
         L     0;
         T     #STC_tPROP.iSyncState;
         L     3;
         T     #OUT_iRetVal;
         BEU;

   e006: A     #STC_tW_MngSysReg.tST.xDone;
         JCN   s006;

         L     6;
         T     #STC_tPROP.iSyncState;

         CALL  FILL
         ( BVAL    := #TMP_dZero,
           RET_VAL := #TMP_iAuxRetVal,
           BLK     := #STC_tW_MngSysReg
         );
         JU    out;
   s006: NOP   0;
END_REGION

REGION Network 9 (STL): RESET "PING" (BIT 1) IN STW1 OF CU
         L     #STC_tPROP.iSyncState;
         L     6;
         ==I;
         JCN   s007;

         SET;
         R     #STC_tPZD_CU.tW.tSTW1.x1;

         L     7;
         T     #STC_tPROP.iSyncState;
         JU    out;
   s007: NOP   0;
END_REGION

REGION Network 10 (STL): SET DONE
         L     #STC_tPROP.iSyncState;
         L     7;
         ==I;
         JCN   s008;

         S     #OUT_xDone;

         L     W#16#0;
         T     #STC_tPROP.iSyncState;

   s008: NOP   0;
END_REGION

REGION Network 11 (STL): Copy Output
   out:  L     #STC_tSYS_DATA.iIOAddress_CU;
         SLW   3;
         T     #TMP_dIO_Pointer;

         L;
         +     48;
         T     #TMP_dPZD_Pointer;

         L     DIW[ #TMP_dPZD_Pointer];
         L     W#16#2;
         AW;
         L     QW[ #TMP_dIO_Pointer];
         OW;
         T     QW[ #TMP_dIO_Pointer];

         BEU;
END_REGION

REGION Network 12 (STL): CU Address wrong
   NWCU: SET;
         S     #OUT_xError;

         L     4;
         T     #OUT_iRetVal;
END_REGION
END_FUNCTION_BLOCK

// folder: 03_Programs_Logics/MCC1201/30_InterfaceEmergencyCutting

FUNCTION_BLOCK "FB_IO_EmergencyCuttingBridge"   // FB28, LAD
{ S7_Optimized_Access := 'TRUE' }
VERSION : 0.1
   VAR_INPUT
      IN_xCycleON : Bool;   // Cycle ON
      IN_xCycleONDel : Bool;   // Delayed cycle ON signal
      IN_xResetAlarms : Bool;   // Reset alarms
      IN_xFaultsEnabled : Bool;   // Faults enabled
      IN_xMachineReady : Bool;   // Machine ready
      IN_xStartCutCycle : Bool;   // StartCutCycle
      IN_xStartCutForBreak : Bool;
      IN_xProtection : Bool;   // EM Xcut protection
      IN_dConvSpeed : DInt;
      IN_xSimulationActive : Bool;
   END_VAR
   VAR_OUTPUT
      OUT_xStartCutCycle : Bool;
      OUT_xSpare : Bool;
      OUT_xSnap : Bool;
      OUT_xAccelaration : Bool;
   END_VAR
   VAR
      ST_xMachineAnomaly : Bool;   // Machine anomaly
      ST_xStoppingFaults : Bool;   // Stopping fault
      ST_xFaults : Bool;   // Fault
      ST_xWarnings : Bool;   // Warnings
      ST_xConditionOkStopCycle : Bool;   // Condition ok stop cycle
      ST_xOutputEnable : Bool;   // Output enable
      ST_xStartcut : Bool;   // Start Cut
      ST_xStartCutForTrak : Bool;
      ST_xRiseAfterDescence : Bool;
      ST_TrackingOnZone_0 : Bool;   // ST_Tracking On Zone0 (0-500)
      ST_TrackingOnZone_1 : Bool;   // ST_Tracking On Zone0 (500-1000)
      ST_TrackingOnZone_2 : Bool;   // ST_Tracking On Zone0 (1000-1500)
      ST_TrackingOnZone_3 : Bool;   // ST_Tracking On Zone0 (1500-2000)
      ST_TrackingOnZone_4 : Bool;   // ST_Tracking On Zone0 (2500-3000)
      ST_TrackingOnZone_5 : Bool;   // ST_Tracking On Zone0 (3500-4000)
      ST_TrackingOnZone_6 : Bool;   // ST_Tracking On Zone0 (3500-4000)
      Os_Ready : Bool;
      Os_Readys : Bool;
      Os_StartCut : Bool;
      OSR_CyclecuttingON : Bool;
      OUTPUT_xMachineRun : Bool;   // Output machine run
      Aux_CountStartCut : Real;
      Aux_trackingcount_0 : Real;
      Aux_trackingCount_1 : Real;
      Aux_trackingCount_2 : Real;
      Aux_trackingCount_3 : Real;
      Aux_trackingCount_4 : Real;
      Aux_trackingCount_5 : Real;
      Aux_trackingCount_6 : Real;
      Aux_supportTargetSnap : Real;
      Aux_supportTargetAcc : Real;
      Aux_AccelerationSpace_mm : Real;
      Aux_dTimeCut : DInt;
      Aux_rSpaceXscan : Real;   // mm done every scan
      StartCutTimerOn : TON_TIME;
      SnapOff : TON_TIME;
      tmON_StartCut : "UDT_IECTON_V1.00";
      tmOFF_AccDelay : TP_TIME;
      tHMR : Struct   // {[Unit]|[Scada Unit]|[LowLimit]|[HigLimit]|[Acces]}
         dState : Int;   // State Conveyor (1=No anomaly, 3=Run, 7=Anomaly) {x|x|x|x|O}
         dDistanceFromSnaproll_cmm : DInt;   // Distance from snaproll [mm/100] {mm/100|mm|0|60000|M}
      END_STRUCT;
      tHMW : Struct   // {[Unit]|[Scada Unit]|[LowLimit]|[HigLimit]|[Acces]}
         rPlateLenght_mm : Real;   // Maximum plate lenght for contrast enabling [mm] {mm|mm|1|7000|O}
         rBreakPosOffset_mm : Real;   // BreakOffset [mm] {mm|mm|1|1000|O}
         dSnapDuration_ms : DInt;   // Time snap in up position [ms] {ms|s|0|1|O}
         dAccelerationDelay_ms : DInt;   // acceleration delay [ms] {ms|s|0|1|O}
         xUpdateDistSnap : Bool;   // Update distance from snap roll {x|x|x|x|M}
         dDistanceFromSnaproll_cmm : DInt;   // Distance from snaproll [mm/100] [mm/100] {mm/100|mm|0|60000|M}
      END_STRUCT;
      tALM : Struct   // HMI Alarms
         tS : Struct   // Stopping faults
            xMachineNotReady : Bool;   // Machine not ready
            xQMProtection : Bool;   // QM Protection
            xSpare_2 : Bool;
            xSpare_3 : Bool;
            xSpare_4 : Bool;
            xSpare_5 : Bool;
            xSpare_6 : Bool;
            xSpare_7 : Bool;
            xSpare_8 : Bool;
            xSpare_9 : Bool;
            xSpare_10 : Bool;
            xSpare_11 : Bool;
            xSpare_12 : Bool;
            xSpare_13 : Bool;
            xSpare_14 : Bool;
            xSpare_15 : Bool;
            xSpare_16 : Bool;
            xSpare_17 : Bool;
            xSpare_18 : Bool;
            xSpare_19 : Bool;
            xSpare_20 : Bool;
            xSpare_21 : Bool;
            xSpare_22 : Bool;
            xSpare_23 : Bool;
            xSpare_24 : Bool;
            xSpare_25 : Bool;
            xSpare_26 : Bool;
            xSpare_27 : Bool;
            xSpare_28 : Bool;
            xSpare_29 : Bool;
            xSpare_30 : Bool;
            xSpare_31 : Bool;
         END_STRUCT;
         tF : Struct   // Faults
            xSpare_0 : Bool;
            xSpare_1 : Bool;
            xSpare_2 : Bool;
            xSpare_3 : Bool;
            xSpare_4 : Bool;
            xSpare_5 : Bool;
            xSpare_6 : Bool;
            xSpare_7 : Bool;
            xSpare_8 : Bool;
            xSpare_9 : Bool;
            xSpare_10 : Bool;
            xSpare_11 : Bool;
            xSpare_12 : Bool;
            xSpare_13 : Bool;
            xSpare_14 : Bool;
            xSpare_15 : Bool;
            xSpare_16 : Bool;
            xSpare_17 : Bool;
            xSpare_18 : Bool;
            xSpare_19 : Bool;
            xSpare_20 : Bool;
            xSpare_21 : Bool;
            xSpare_22 : Bool;
            xSpare_23 : Bool;
            xSpare_24 : Bool;
            xSpare_25 : Bool;
            xSpare_26 : Bool;
            xSpare_27 : Bool;
            xSpare_28 : Bool;
            xSpare_29 : Bool;
            xSpare_30 : Bool;
            xSpare_31 : Bool;
         END_STRUCT;
         tW : Struct   // Warnings
            xSpare_0 : Bool;
            xSpare_1 : Bool;
            xSpare_2 : Bool;
            xSpare_3 : Bool;
            xSpare_4 : Bool;
            xSpare_5 : Bool;
            xSpare_6 : Bool;
            xSpare_7 : Bool;
            xSpare_8 : Bool;
            xSpare_9 : Bool;
            xSpare_10 : Bool;
            xSpare_11 : Bool;
            xSpare_12 : Bool;
            xSpare_13 : Bool;
            xSpare_14 : Bool;
            xSpare_15 : Bool;
            xSpare_16 : Bool;
            xSpare_17 : Bool;
            xSpare_18 : Bool;
            xSpare_19 : Bool;
            xSpare_20 : Bool;
            xSpare_21 : Bool;
            xSpare_22 : Bool;
            xSpare_23 : Bool;
            xSpare_24 : Bool;
            xSpare_25 : Bool;
            xSpare_26 : Bool;
            xSpare_27 : Bool;
            xSpare_28 : Bool;
            xSpare_29 : Bool;
            xSpare_30 : Bool;
            xSpare_31 : Bool;
         END_STRUCT;
      END_STRUCT;
   END_VAR
   VAR_TEMP
      TMP_xDummybit : Bool;
      Tmp_StartCutBreak : Bool;
      TMP_dIndex : DInt;
      TMP_dwValue : DWord;
      TMP_iRetVal : Int;
      Tmp_rSpeed : Real;
      Tmp_rTimeObScan : Real;
   END_VAR
   VAR CONSTANT
      CONST_DBREAKDOWNOFF_CMM : DInt := 100000;   // Break downstream offset [mm/100]
      CONST_DBREAKUPOFF_CMM : DInt := 100000;   // Break upstream offset [mm/100]
   END_VAR
   VAR_TEMP   // added for the SCL form of the ladder/FBD networks
      _w1 : Bool;
      _w2 : Bool;
   END_VAR
BEGIN

REGION Network 1: #####_MATCH_#####
END_REGION

REGION Network 2 (SCL): Simulation
   IF #IN_xSimulationActive THEN
       #IN_xProtection := 1;
       #IN_xMachineReady := 1;
   END_IF;
END_REGION

REGION Network 3: ####_ALARMS_####
END_REGION

REGION Network 4 (SCL): Reset alarms
   IF #IN_xResetAlarms THEN

       #TMP_dwValue := 0;

       SCATTER(IN:=#TMP_dwValue,
               OUT=>#tALM.tS);

       SCATTER(IN:=#TMP_dwValue,
               OUT=>#tALM.tF);

       SCATTER(IN:=#TMP_dwValue,
               OUT=>#tALM.tW);


   END_IF;
END_REGION

REGION Network 5: Local Safety Switch
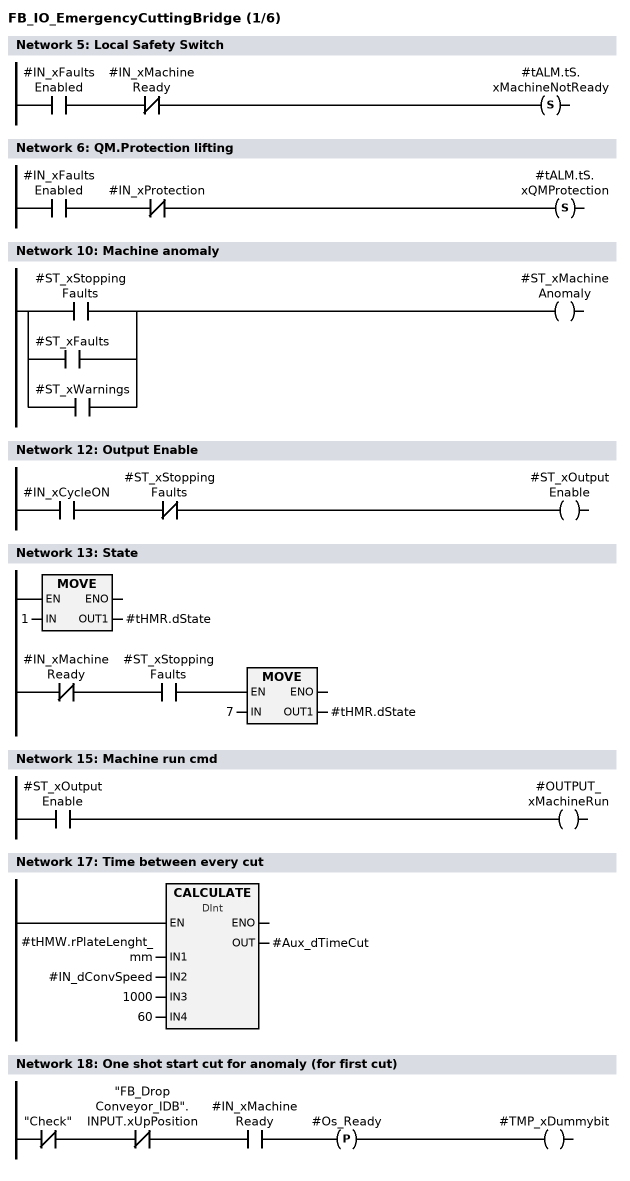
   RUNG wire#powerrail
      Contact( #IN_xFaultsEnabled )
      I_Contact( #IN_xMachineReady )
      S_Coil( #tALM.tS.xMachineNotReady )
   END_RUNG
   // the same network as SCL:
   IF #IN_xFaultsEnabled AND NOT #IN_xMachineReady THEN #tALM.tS.xMachineNotReady := TRUE; END_IF;
END_REGION

REGION Network 6: QM.Protection lifting
   RUNG wire#powerrail
      Contact( #IN_xFaultsEnabled )
      I_Contact( #IN_xProtection )
      S_Coil( #tALM.tS.xQMProtection )
   END_RUNG
   // the same network as SCL:
   IF #IN_xFaultsEnabled AND NOT #IN_xProtection THEN #tALM.tS.xQMProtection := TRUE; END_IF;
END_REGION

REGION Network 7 (SCL): Calculate general statuses
   GATHER(IN:=#tALM.tS,
          OUT=>#TMP_dwValue);

   IF #TMP_dwValue <> 0 THEN
       #ST_xStoppingFaults := TRUE;
   ELSE
       #ST_xStoppingFaults := FALSE;
   END_IF;

   GATHER(IN:=#tALM.tF,
          OUT=>#TMP_dwValue);

   IF #TMP_dwValue <> 0 THEN
       #ST_xFaults := TRUE;
   ELSE
       #ST_xFaults := FALSE;
   END_IF;

   GATHER(IN:=#tALM.tW,
          OUT=>#TMP_dwValue);

   IF #TMP_dwValue <> 0 THEN
       #ST_xWarnings := TRUE;
   ELSE
       #ST_xWarnings := FALSE;
   END_IF;
END_REGION

REGION Network 8 (SCL): Check glass break on Emergency Xcut M203
   "DB_RibbonData".rgtGlassBreakRequest["DGLASSBREAKGET_M203"].IN_dDistanceSnaproll_cmm :=#tHMR.dDistanceFromSnaproll_cmm;
   "DB_RibbonData".rgtGlassBreakRequest["DGLASSBREAKGET_M203"].IN_dDownstreamOffset_cmm := #CONST_DBREAKDOWNOFF_CMM;
   "DB_RibbonData".rgtGlassBreakRequest["DGLASSBREAKGET_M203"].IN_dUpstreamOffset_cmm := #CONST_DBREAKUPOFF_CMM;

   IF "DB_RibbonData".rgtGlassBreakRequest["DGLASSBREAKGET_M203"].OUT_xDataReady THEN
       "Z200".ST_xM203GlassBreak := "DB_RibbonData".rgtGlassBreakRequest["DGLASSBREAKGET_M203"].OUT_xGlassBreak;
   END_IF;

   IF "DB_RibbonData".rgtGlassBreakRequest["DGLASSBREAKGET_M203"].OUT_xDataReady OR NOT "DB_RibbonData".rgtGlassBreakRequest["DGLASSBREAKGET_M203"].IN_xRequestGlassBreak THEN
       "DB_RibbonData".rgtGlassBreakRequest["DGLASSBREAKGET_M203"].OUT_xDataReady := FALSE;
       "DB_RibbonData".rgtGlassBreakRequest["DGLASSBREAKGET_M203"].IN_xRequestGlassBreak := TRUE;
   END_IF;
END_REGION

REGION Network 9: #####_HMI_LOGICS_#####
END_REGION

REGION Network 10: Machine anomaly
   RUNG wire#powerrail
      Contact( #ST_xStoppingFaults )
      wire#w1
      Coil( #ST_xMachineAnomaly )
   END_RUNG
   RUNG wire#powerrail
      Contact( #ST_xFaults )
   END_RUNG wire#w1
   RUNG wire#powerrail
      Contact( #ST_xWarnings )
   END_RUNG wire#w1
   // the same network as SCL:
   #ST_xMachineAnomaly := #ST_xStoppingFaults OR #ST_xFaults OR #ST_xWarnings;
END_REGION

REGION Network 11 (SCL): Distance from snap roll EM Xcut
   REGION UpdateDistanceSnaproll

   IF #tHMW.xUpdateDistSnap THEN
       #tHMW.xUpdateDistSnap := FALSE;

       #tHMR.dDistanceFromSnaproll_cmm := #tHMW.dDistanceFromSnaproll_cmm;

   END_IF;

   END_REGION
END_REGION

REGION Network 12: Output Enable
   RUNG wire#powerrail
      Contact( #IN_xCycleON )
      I_Contact( #ST_xStoppingFaults )
      Coil( #ST_xOutputEnable )
   END_RUNG
   // the same network as SCL:
   #ST_xOutputEnable := #IN_xCycleON AND NOT #ST_xStoppingFaults;
END_REGION

REGION Network 13: State
   RUNG wire#powerrail
      Move(in := 1, out1 => #tHMR.dState)
   END_RUNG
   RUNG wire#powerrail
      I_Contact( #IN_xMachineReady )
      Contact( #ST_xStoppingFaults )
      Move(in := 7, out1 => #tHMR.dState)
   END_RUNG
   // the same network as SCL:
   #tHMR.dState := 1;
   IF NOT #IN_xMachineReady AND #ST_xStoppingFaults THEN #tHMR.dState := 7; END_IF;
END_REGION

REGION Network 14: #####_OUTPUT_#####
END_REGION

REGION Network 15: Machine run cmd
   RUNG wire#powerrail
      Contact( #ST_xOutputEnable )
      Coil( #OUTPUT_xMachineRun )
   END_RUNG
   // the same network as SCL:
   #OUTPUT_xMachineRun := #ST_xOutputEnable;
END_REGION

REGION Network 16 (SCL): Space[mm] done in 10 ms
   #Tmp_rSpeed :=   DINT_TO_REAL (#IN_dConvSpeed) ;

   #Aux_rSpaceXscan := ((#Tmp_rSpeed / 60.0) / 1000.0) * "GP_OB_Initialize_Main_IDB".OUT_dExecutionTime_ms;
END_REGION

REGION Network 17: Time between every cut
   RUNG wire#powerrail
      { S7_Templates := "SrcType := DInt"; S7_Expression := "(IN1*IN3)/(IN2/IN4)" } Calculate(in1 := #tHMW.rPlateLenght_mm, in2 := #IN_dConvSpeed, in3 := 1000, in4 := 60, out => #Aux_dTimeCut)
   END_RUNG
   // the same network as SCL:
   #Aux_dTimeCut := (#tHMW.rPlateLenght_mm*1000)/(#IN_dConvSpeed/60);
END_REGION

REGION Network 18: One shot start cut for anomaly (for first cut)
   RUNG wire#powerrail
      I_Contact( "Check" )
      I_Contact( "FB_DropConveyor_IDB".INPUT.xUpPosition )
      Contact( #IN_xMachineReady )
      P_Trig( #Os_Ready )
      Coil( #TMP_xDummybit )
   END_RUNG
   // the same network as SCL:
   #_w1 := NOT "Check" AND NOT "FB_DropConveyor_IDB".INPUT.xUpPosition AND #IN_xMachineReady;
   #_w2 := #_w1 AND NOT #Os_Ready;   // rising edge
   #Os_Ready := #_w1;
   #TMP_xDummybit := #_w2;
END_REGION

REGION Network 19: Start cut for tracking
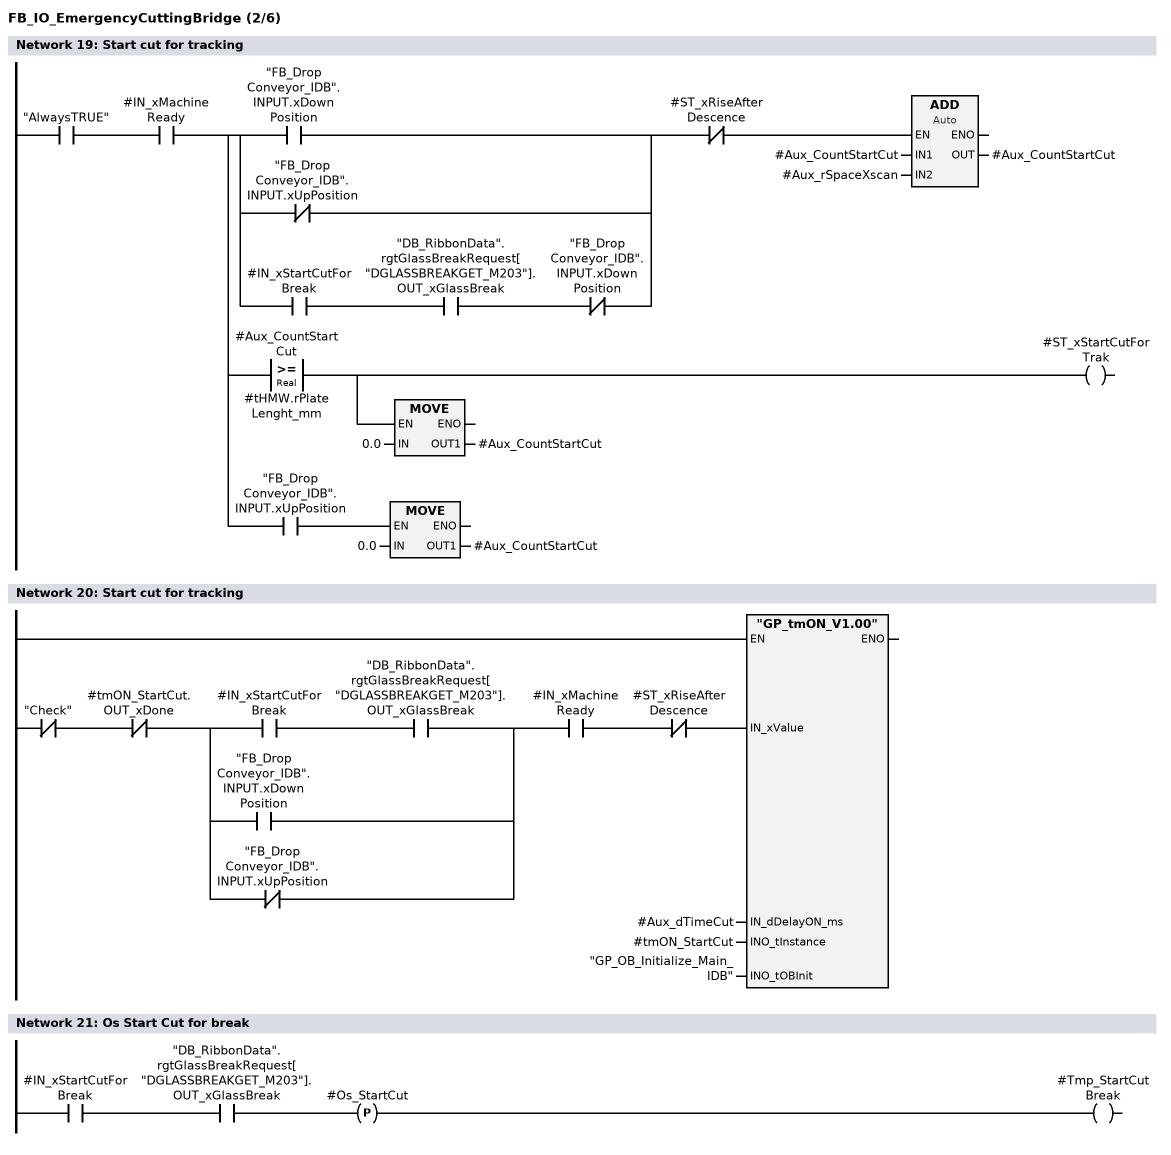
   RUNG wire#powerrail
      Contact( "AlwaysTRUE" )
      Contact( #IN_xMachineReady )
      wire#w1
      Contact( "FB_DropConveyor_IDB".INPUT.xDownPosition )
      wire#w2
      I_Contact( #ST_xRiseAfterDescence )
      Add(in1 := #Aux_CountStartCut, in2 := #Aux_rSpaceXscan, out => #Aux_CountStartCut)
   END_RUNG
   RUNG wire#w1
      I_Contact( "FB_DropConveyor_IDB".INPUT.xUpPosition )
   END_RUNG wire#w2
   RUNG wire#w1
      Contact( #IN_xStartCutForBreak )
      Contact( "DB_RibbonData".rgtGlassBreakRequest["DGLASSBREAKGET_M203"].OUT_xGlassBreak )
      I_Contact( "FB_DropConveyor_IDB".INPUT.xDownPosition )
   END_RUNG wire#w2
   RUNG wire#w1
      { S7_Templates := "SrcType := Real" } GE_Contact(in1 := #Aux_CountStartCut, in2 := #tHMW.rPlateLenght_mm)
      wire#w3
      Coil( #ST_xStartCutForTrak )
   END_RUNG
   RUNG wire#w3
      Move(in := 0.0, out1 => #Aux_CountStartCut)
   END_RUNG
   RUNG wire#w1
      Contact( "FB_DropConveyor_IDB".INPUT.xUpPosition )
      Move(in := 0.0, out1 => #Aux_CountStartCut)
   END_RUNG
   // the same network as SCL:
   #_w1 := "AlwaysTRUE" AND #IN_xMachineReady;
   IF #_w1 AND ("FB_DropConveyor_IDB".INPUT.xDownPosition OR NOT "FB_DropConveyor_IDB".INPUT.xUpPosition OR (#IN_xStartCutForBreak AND "DB_RibbonData".rgtGlassBreakRequest["DGLASSBREAKGET_M203"].OUT_xGlassBreak AND NOT "FB_DropConveyor_IDB".INPUT.xDownPosition)) AND NOT #ST_xRiseAfterDescence THEN
       #Aux_CountStartCut := #Aux_CountStartCut + #Aux_rSpaceXscan;
   END_IF;
   #ST_xStartCutForTrak := #_w1 AND (#Aux_CountStartCut >= #tHMW.rPlateLenght_mm);
   IF #ST_xStartCutForTrak THEN #Aux_CountStartCut := 0.0; END_IF;
   IF #_w1 AND "FB_DropConveyor_IDB".INPUT.xUpPosition THEN #Aux_CountStartCut := 0.0; END_IF;
END_REGION

REGION Network 20: Start cut for tracking
   RUNG wire#powerrail
      "GP_tmON_V1.00"(IN_xValue := wire#w3, IN_dDelayON_ms := #Aux_dTimeCut, INO_tInstance := #tmON_StartCut, INO_tOBInit := "GP_OB_Initialize_Main_IDB")
   END_RUNG
   RUNG wire#powerrail
      I_Contact( "Check" )
      I_Contact( #tmON_StartCut.OUT_xDone )
      wire#w1
      Contact( #IN_xStartCutForBreak )
      Contact( "DB_RibbonData".rgtGlassBreakRequest["DGLASSBREAKGET_M203"].OUT_xGlassBreak )
      wire#w2
      Contact( #IN_xMachineReady )
      I_Contact( #ST_xRiseAfterDescence )
   END_RUNG wire#w3
   RUNG wire#w1
      Contact( "FB_DropConveyor_IDB".INPUT.xDownPosition )
   END_RUNG wire#w2
   RUNG wire#w1
      I_Contact( "FB_DropConveyor_IDB".INPUT.xUpPosition )
   END_RUNG wire#w2
   // the same network as SCL:
   "GP_tmON_V1.00"(IN_xValue := NOT "Check" AND NOT #tmON_StartCut.OUT_xDone AND ((#IN_xStartCutForBreak AND "DB_RibbonData".rgtGlassBreakRequest["DGLASSBREAKGET_M203"].OUT_xGlassBreak) OR "FB_DropConveyor_IDB".INPUT.xDownPosition OR NOT "FB_DropConveyor_IDB".INPUT.xUpPosition) AND #IN_xMachineReady AND NOT #ST_xRiseAfterDescence,
                   IN_dDelayON_ms := #Aux_dTimeCut,
                   INO_tInstance := #tmON_StartCut,
                   INO_tOBInit := "GP_OB_Initialize_Main_IDB");
END_REGION

REGION Network 21: Os Start Cut for break
   RUNG wire#powerrail
      Contact( #IN_xStartCutForBreak )
      Contact( "DB_RibbonData".rgtGlassBreakRequest["DGLASSBREAKGET_M203"].OUT_xGlassBreak )
      P_Trig( #Os_StartCut )
      Coil( #Tmp_StartCutBreak )
   END_RUNG
   // the same network as SCL:
   #_w1 := #IN_xStartCutForBreak AND "DB_RibbonData".rgtGlassBreakRequest["DGLASSBREAKGET_M203"].OUT_xGlassBreak;
   #_w2 := #_w1 AND NOT #Os_StartCut;   // rising edge
   #Os_StartCut := #_w1;
   #Tmp_StartCutBreak := #_w2;
END_REGION

REGION Network 22: Start Cut
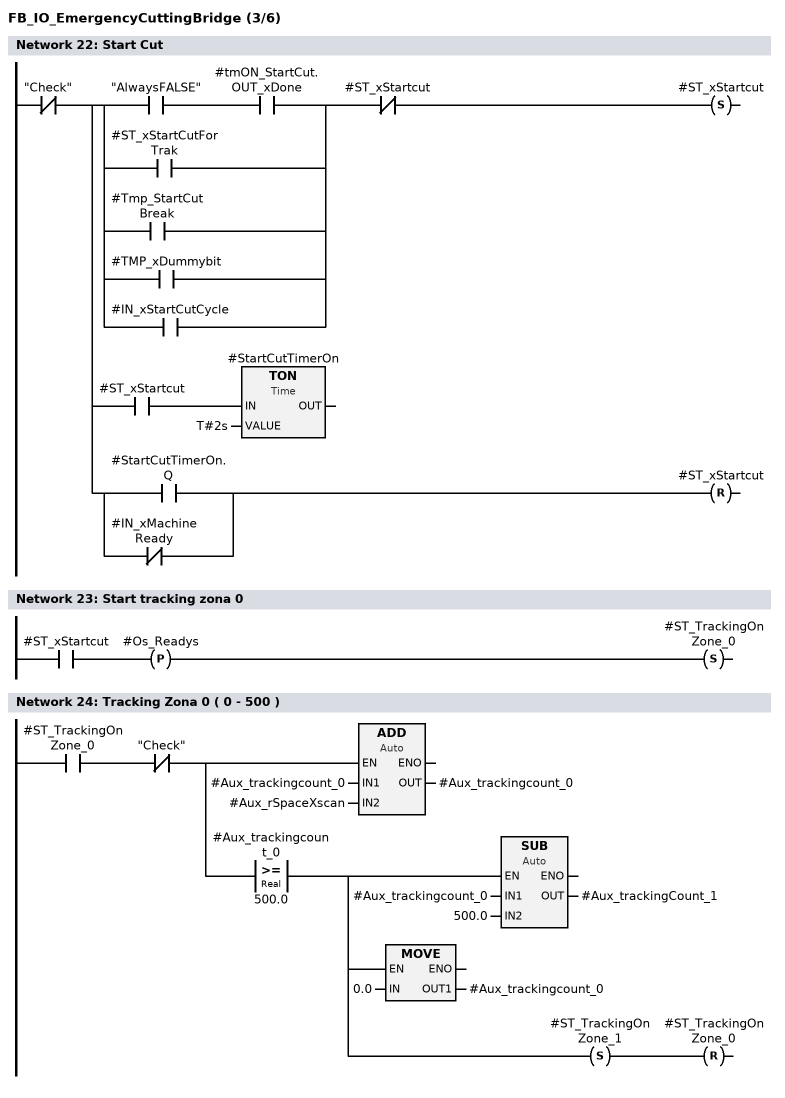
   IF NOT "Check" AND (("AlwaysFALSE" AND #tmON_StartCut.OUT_xDone) OR #ST_xStartCutForTrak OR #Tmp_StartCutBreak OR #TMP_xDummybit OR #IN_xStartCutCycle) AND NOT #ST_xStartcut THEN
       #ST_xStartcut := TRUE;
   END_IF;
   #StartCutTimerOn(IN := NOT "Check" AND #ST_xStartcut, PT := T#2s);   // TON coil
   IF NOT "Check" AND (#StartCutTimerOn.Q OR NOT #IN_xMachineReady) THEN #ST_xStartcut := FALSE; END_IF;
END_REGION

REGION Network 23: Start tracking zona 0
   RUNG wire#powerrail
      Contact( #ST_xStartcut )
      P_Trig( #Os_Readys )
      S_Coil( #ST_TrackingOnZone_0 )
   END_RUNG
   // the same network as SCL:
   #_w1 := #ST_xStartcut AND NOT #Os_Readys;   // rising edge
   #Os_Readys := #ST_xStartcut;
   IF #_w1 THEN #ST_TrackingOnZone_0 := TRUE; END_IF;
END_REGION

REGION Network 24: Tracking Zona 0 ( 0 - 500 )
   RUNG wire#powerrail
      Contact( #ST_TrackingOnZone_0 )
      I_Contact( "Check" )
      wire#w1
      Add(in1 := #Aux_trackingcount_0, in2 := #Aux_rSpaceXscan, out => #Aux_trackingcount_0)
   END_RUNG
   RUNG wire#w1
      { S7_Templates := "SrcType := Real" } GE_Contact(in1 := #Aux_trackingcount_0, in2 := 500.0)
      wire#w2
      Sub(in1 := #Aux_trackingcount_0, in2 := 500.0, out => #Aux_trackingCount_1)
   END_RUNG
   RUNG wire#w2
      Move(in := 0.0, out1 => #Aux_trackingcount_0)
   END_RUNG
   RUNG wire#w2
      S_Coil( #ST_TrackingOnZone_1 )
      R_Coil( #ST_TrackingOnZone_0 )
   END_RUNG
   // the same network as SCL:
   #_w1 := #ST_TrackingOnZone_0 AND NOT "Check";
   IF #_w1 THEN #Aux_trackingcount_0 := #Aux_trackingcount_0 + #Aux_rSpaceXscan; END_IF;
   IF #_w1 AND (#Aux_trackingcount_0 >= 500.0) THEN
       #Aux_trackingCount_1 := #Aux_trackingcount_0 - 500.0;
   END_IF;
   #_w2 := #_w1 AND (#Aux_trackingcount_0 >= 500.0);
   IF #_w2 THEN
       #Aux_trackingcount_0 := 0.0;
       #ST_TrackingOnZone_1 := TRUE;
       #ST_TrackingOnZone_0 := FALSE;
   END_IF;
END_REGION

REGION Network 25: Tracking Zona 1 ( 500-1000 )
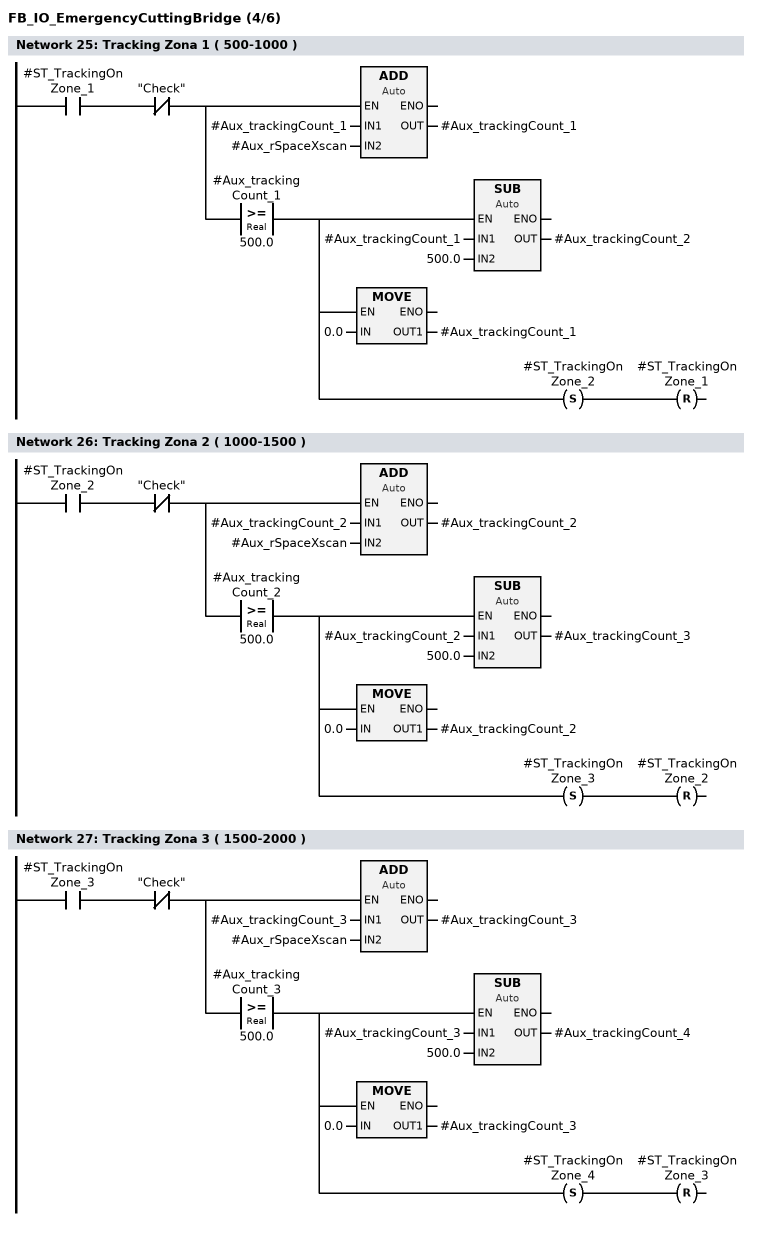
   RUNG wire#powerrail
      Contact( #ST_TrackingOnZone_1 )
      I_Contact( "Check" )
      wire#w1
      Add(in1 := #Aux_trackingCount_1, in2 := #Aux_rSpaceXscan, out => #Aux_trackingCount_1)
   END_RUNG
   RUNG wire#w1
      { S7_Templates := "SrcType := Real" } GE_Contact(in1 := #Aux_trackingCount_1, in2 := 500.0)
      wire#w2
      Sub(in1 := #Aux_trackingCount_1, in2 := 500.0, out => #Aux_trackingCount_2)
   END_RUNG
   RUNG wire#w2
      Move(in := 0.0, out1 => #Aux_trackingCount_1)
   END_RUNG
   RUNG wire#w2
      S_Coil( #ST_TrackingOnZone_2 )
      R_Coil( #ST_TrackingOnZone_1 )
   END_RUNG
   // the same network as SCL:
   #_w1 := #ST_TrackingOnZone_1 AND NOT "Check";
   IF #_w1 THEN #Aux_trackingCount_1 := #Aux_trackingCount_1 + #Aux_rSpaceXscan; END_IF;
   IF #_w1 AND (#Aux_trackingCount_1 >= 500.0) THEN
       #Aux_trackingCount_2 := #Aux_trackingCount_1 - 500.0;
   END_IF;
   #_w2 := #_w1 AND (#Aux_trackingCount_1 >= 500.0);
   IF #_w2 THEN
       #Aux_trackingCount_1 := 0.0;
       #ST_TrackingOnZone_2 := TRUE;
       #ST_TrackingOnZone_1 := FALSE;
   END_IF;
END_REGION

REGION Network 26: Tracking Zona 2 ( 1000-1500 )
   RUNG wire#powerrail
      Contact( #ST_TrackingOnZone_2 )
      I_Contact( "Check" )
      wire#w1
      Add(in1 := #Aux_trackingCount_2, in2 := #Aux_rSpaceXscan, out => #Aux_trackingCount_2)
   END_RUNG
   RUNG wire#w1
      { S7_Templates := "SrcType := Real" } GE_Contact(in1 := #Aux_trackingCount_2, in2 := 500.0)
      wire#w2
      Sub(in1 := #Aux_trackingCount_2, in2 := 500.0, out => #Aux_trackingCount_3)
   END_RUNG
   RUNG wire#w2
      Move(in := 0.0, out1 => #Aux_trackingCount_2)
   END_RUNG
   RUNG wire#w2
      S_Coil( #ST_TrackingOnZone_3 )
      R_Coil( #ST_TrackingOnZone_2 )
   END_RUNG
   // the same network as SCL:
   #_w1 := #ST_TrackingOnZone_2 AND NOT "Check";
   IF #_w1 THEN #Aux_trackingCount_2 := #Aux_trackingCount_2 + #Aux_rSpaceXscan; END_IF;
   IF #_w1 AND (#Aux_trackingCount_2 >= 500.0) THEN
       #Aux_trackingCount_3 := #Aux_trackingCount_2 - 500.0;
   END_IF;
   #_w2 := #_w1 AND (#Aux_trackingCount_2 >= 500.0);
   IF #_w2 THEN
       #Aux_trackingCount_2 := 0.0;
       #ST_TrackingOnZone_3 := TRUE;
       #ST_TrackingOnZone_2 := FALSE;
   END_IF;
END_REGION

REGION Network 27: Tracking Zona 3 ( 1500-2000 )
   RUNG wire#powerrail
      Contact( #ST_TrackingOnZone_3 )
      I_Contact( "Check" )
      wire#w1
      Add(in1 := #Aux_trackingCount_3, in2 := #Aux_rSpaceXscan, out => #Aux_trackingCount_3)
   END_RUNG
   RUNG wire#w1
      { S7_Templates := "SrcType := Real" } GE_Contact(in1 := #Aux_trackingCount_3, in2 := 500.0)
      wire#w2
      Sub(in1 := #Aux_trackingCount_3, in2 := 500.0, out => #Aux_trackingCount_4)
   END_RUNG
   RUNG wire#w2
      Move(in := 0.0, out1 => #Aux_trackingCount_3)
   END_RUNG
   RUNG wire#w2
      S_Coil( #ST_TrackingOnZone_4 )
      R_Coil( #ST_TrackingOnZone_3 )
   END_RUNG
   // the same network as SCL:
   #_w1 := #ST_TrackingOnZone_3 AND NOT "Check";
   IF #_w1 THEN #Aux_trackingCount_3 := #Aux_trackingCount_3 + #Aux_rSpaceXscan; END_IF;
   IF #_w1 AND (#Aux_trackingCount_3 >= 500.0) THEN
       #Aux_trackingCount_4 := #Aux_trackingCount_3 - 500.0;
   END_IF;
   #_w2 := #_w1 AND (#Aux_trackingCount_3 >= 500.0);
   IF #_w2 THEN
       #Aux_trackingCount_3 := 0.0;
       #ST_TrackingOnZone_4 := TRUE;
       #ST_TrackingOnZone_3 := FALSE;
   END_IF;
END_REGION

REGION Network 28: Tracking Zona 4 ( 2000-2500 )
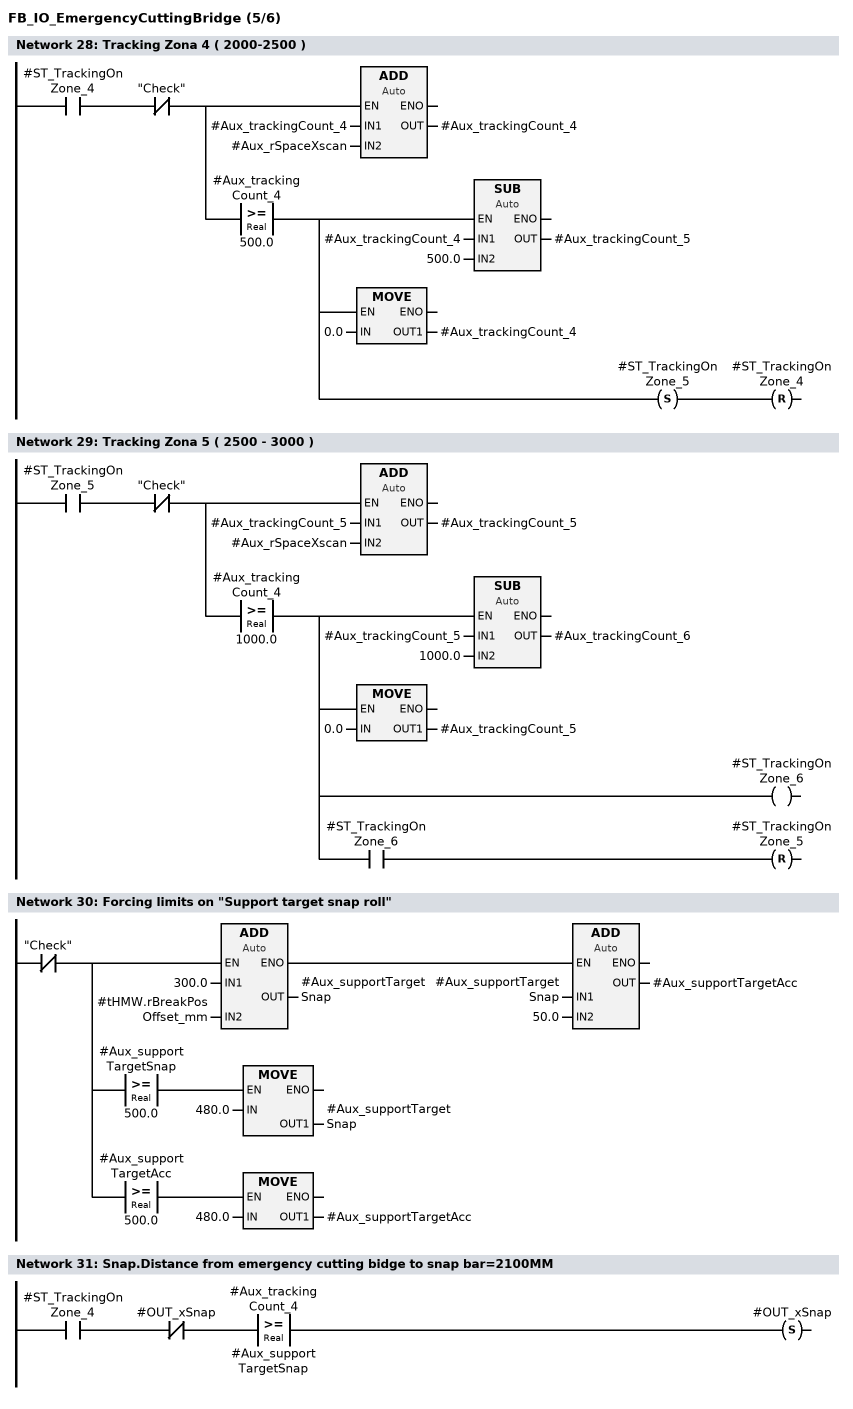
   RUNG wire#powerrail
      Contact( #ST_TrackingOnZone_4 )
      I_Contact( "Check" )
      wire#w1
      Add(in1 := #Aux_trackingCount_4, in2 := #Aux_rSpaceXscan, out => #Aux_trackingCount_4)
   END_RUNG
   RUNG wire#w1
      { S7_Templates := "SrcType := Real" } GE_Contact(in1 := #Aux_trackingCount_4, in2 := 500.0)
      wire#w2
      Sub(in1 := #Aux_trackingCount_4, in2 := 500.0, out => #Aux_trackingCount_5)
   END_RUNG
   RUNG wire#w2
      Move(in := 0.0, out1 => #Aux_trackingCount_4)
   END_RUNG
   RUNG wire#w2
      S_Coil( #ST_TrackingOnZone_5 )
      R_Coil( #ST_TrackingOnZone_4 )
   END_RUNG
   // the same network as SCL:
   #_w1 := #ST_TrackingOnZone_4 AND NOT "Check";
   IF #_w1 THEN #Aux_trackingCount_4 := #Aux_trackingCount_4 + #Aux_rSpaceXscan; END_IF;
   IF #_w1 AND (#Aux_trackingCount_4 >= 500.0) THEN
       #Aux_trackingCount_5 := #Aux_trackingCount_4 - 500.0;
   END_IF;
   #_w2 := #_w1 AND (#Aux_trackingCount_4 >= 500.0);
   IF #_w2 THEN
       #Aux_trackingCount_4 := 0.0;
       #ST_TrackingOnZone_5 := TRUE;
       #ST_TrackingOnZone_4 := FALSE;
   END_IF;
END_REGION

REGION Network 29: Tracking Zona 5 ( 2500 - 3000 )
   RUNG wire#powerrail
      Contact( #ST_TrackingOnZone_5 )
      I_Contact( "Check" )
      wire#w1
      Add(in1 := #Aux_trackingCount_5, in2 := #Aux_rSpaceXscan, out => #Aux_trackingCount_5)
   END_RUNG
   RUNG wire#w1
      { S7_Templates := "SrcType := Real" } GE_Contact(in1 := #Aux_trackingCount_4, in2 := 1000.0)
      wire#w2
      Sub(in1 := #Aux_trackingCount_5, in2 := 1000.0, out => #Aux_trackingCount_6)
   END_RUNG
   RUNG wire#w2
      Move(in := 0.0, out1 => #Aux_trackingCount_5)
   END_RUNG
   RUNG wire#w2
      Coil( #ST_TrackingOnZone_6 )
   END_RUNG
   RUNG wire#w2
      Contact( #ST_TrackingOnZone_6 )
      R_Coil( #ST_TrackingOnZone_5 )
   END_RUNG
   // the same network as SCL:
   #_w1 := #ST_TrackingOnZone_5 AND NOT "Check";
   IF #_w1 THEN #Aux_trackingCount_5 := #Aux_trackingCount_5 + #Aux_rSpaceXscan; END_IF;
   #_w2 := #_w1 AND (#Aux_trackingCount_4 >= 1000.0);
   IF #_w2 THEN
       #Aux_trackingCount_6 := #Aux_trackingCount_5 - 1000.0;
       #Aux_trackingCount_5 := 0.0;
   END_IF;
   #ST_TrackingOnZone_6 := #_w2;
   IF #_w2 AND #ST_TrackingOnZone_6 THEN #ST_TrackingOnZone_5 := FALSE; END_IF;
END_REGION

REGION Network 30: Forcing limits on "Support target snap roll"
   RUNG wire#powerrail
      I_Contact( "Check" )
      wire#w1
      Add(in1 := 300.0, in2 := #tHMW.rBreakPosOffset_mm, out => #Aux_supportTargetSnap)
      Add(in1 := #Aux_supportTargetSnap, in2 := 50.0, out => #Aux_supportTargetAcc)
   END_RUNG
   RUNG wire#w1
      { S7_Templates := "SrcType := Real" } GE_Contact(in1 := #Aux_supportTargetSnap, in2 := 500.0)
      Move(in := 480.0, out1 => #Aux_supportTargetSnap)
   END_RUNG
   RUNG wire#w1
      { S7_Templates := "SrcType := Real" } GE_Contact(in1 := #Aux_supportTargetAcc, in2 := 500.0)
      Move(in := 480.0, out1 => #Aux_supportTargetAcc)
   END_RUNG
   // the same network as SCL:
   IF NOT "Check" THEN
       #Aux_supportTargetSnap := 300.0 + #tHMW.rBreakPosOffset_mm;
       #Aux_supportTargetAcc := #Aux_supportTargetSnap + 50.0;
   END_IF;
   IF NOT "Check" AND (#Aux_supportTargetSnap >= 500.0) THEN #Aux_supportTargetSnap := 480.0; END_IF;
   IF NOT "Check" AND (#Aux_supportTargetAcc >= 500.0) THEN #Aux_supportTargetAcc := 480.0; END_IF;
END_REGION

REGION Network 31: Snap.Distance from emergency cutting bidge to snap bar=2100MM
   RUNG wire#powerrail
      Contact( #ST_TrackingOnZone_4 )
      I_Contact( #OUT_xSnap )
      { S7_Templates := "SrcType := Real" } GE_Contact(in1 := #Aux_trackingCount_4, in2 := #Aux_supportTargetSnap)
      S_Coil( #OUT_xSnap )
   END_RUNG
   // the same network as SCL:
   IF #ST_TrackingOnZone_4 AND NOT #OUT_xSnap AND (#Aux_trackingCount_4 >= #Aux_supportTargetSnap) THEN
       #OUT_xSnap := TRUE;
   END_IF;
END_REGION

REGION Network 32: snap duration